   N233 : DINT[1] := ([0] := 9);
   N24 : DINT[31] := ([0] := 100, [1] := 1, [2] := 100, [3] := 1, [4] := 5, [5] := 5, [6] := 60, [7] := 1, [8] := 100, [9] := 1, [10] := 100, [11] := 1, [12] := 5, [13] := 5, [14] := 60, [15] := 1);
   N240 : DINT[68] := ([8] := 254, [10] := -256, [50] := 128, [51] := 9, [52] := 210, [54] := 1, [55] := 210, [60] := 25600, [61] := 9, [62] := 210, [64] := 17408, [66] := 210);
   N241 : DINT[1];
   N242 : DINT[2] := ([0] := -9, [1] := -9);
   N250 : DINT[100] := ([8] := 99, [10] := -256, [50] := -32640, [51] := 9, [52] := 200, [54] := 1, [55] := 200, [61] := 9, [62] := 200, [65] := 1, [66] := 200);
   N251 : DINT[100];
   N252 : DINT[100] := ([0] := -9, [1] := -9);
   N26 : DINT[33] := ([1] := 8, [10] := 38, [11] := 1, [30] := -15194, [31] := 8);
   N27 : DINT[50] := ([40] := 28176, [41] := 29344, [42] := 23976, [43] := 25960, [44] := 29304, [45] := 27664, [46] := 28928, [47] := 16);
   N28 : DINT[17] := ([0] := 124, [1] := 158, [2] := 937, [3] := 50, [4] := 9, [5] := 156, [6] := 3, [10] := 1000, [12] := 100);
   N7 : DINT[100] := ([0] := 5, [1] := 20, [2] := 20, [4] := 30000, [7] := 48, [8] := 48, [9] := 48, [10] := 53, [11] := 53, [12] := 43, [13] := 46, [14] := 46, [15] := 46, [16] := 51, [17] := 51, [18] := 46, [50] := 1, [51] := 1, [52] := 1, [53] := 1, [54] := 1, [55] := 1, [56] := 1, [57] := 1, [58] := 1, [59] := 1, [60] := 1, [61] := 1, [62] := 1, [93] := 9, [99] := 9);
   N_RECVING_PIT_GATE_AUTO : ALIAS FOR Local:0:I.Data.2;
   N_RECVING_PIT_GATE_CLOSE : ALIAS FOR Local:5:O.Data.5;
   N_RECVING_PIT_GATE_OPEN : ALIAS FOR Local:5:O.Data.4;
   NU : DINT;
   O10 : ALIAS FOR R1S0_AENTR:10:O.Data;
   O10_000_Bit00 : ALIAS FOR O10.0;
   O10_000_Bit01 : ALIAS FOR O10.1;
   O10_000_Bit02 : ALIAS FOR O10.2;
   O10_000_Bit03 : ALIAS FOR O10.3;
   O10_000_Bit04 : ALIAS FOR O10.4;
   O10_000_Bit05 : ALIAS FOR O10.5;
   O10_000_Bit06 : ALIAS FOR O10.6;
   O10_000_Bit07 : ALIAS FOR O10.7;
   O10_000_Bit08 : ALIAS FOR O10.8;
   O10_000_Bit09 : ALIAS FOR O10.9;
   O10_000_Bit10 : ALIAS FOR O10.10;
   O10_000_Bit11 : ALIAS FOR O10.11;
   O10_000_Bit12 : ALIAS FOR O10.12;
   O10_000_Bit13 : ALIAS FOR O10.13;
   O10_000_Bit14 : ALIAS FOR O10.14;
   O10_000_Bit15 : ALIAS FOR O10.15;
   O11 : ALIAS FOR R1S0_AENTR:11:O.Data;
   O11_000_Bit00 : ALIAS FOR O11.0;
   O11_000_Bit01 : ALIAS FOR O11.1;
   O11_000_Bit02 : ALIAS FOR O11.2;
   O11_000_Bit03 : ALIAS FOR O11.3;
   O11_000_Bit04 : ALIAS FOR O11.4;
   O11_000_Bit05 : ALIAS FOR O11.5;
   O11_000_Bit06 : ALIAS FOR O11.6;
   O11_000_Bit07 : ALIAS FOR O11.7;
   O11_000_Bit08 : ALIAS FOR O11.8;
   O11_000_Bit09 : ALIAS FOR O11.9;
   O11_000_Bit10 : ALIAS FOR O11.10;
   O11_000_Bit11 : ALIAS FOR O11.11;
   O11_000_Bit12 : ALIAS FOR O11.12;
   O11_000_Bit13 : ALIAS FOR O11.13;
   O11_000_Bit14 : ALIAS FOR O11.14;
   O12 : ALIAS FOR R1S0_AENTR:12:O.Data;
   O12_000_Bit00 : ALIAS FOR O12.0;
   O12_000_Bit01 : ALIAS FOR O12.1;
   O12_000_Bit02 : ALIAS FOR O12.2;
   O12_000_Bit03 : ALIAS FOR O12.3;
   O12_000_Bit04 : ALIAS FOR O12.4;
   O12_000_Bit05 : ALIAS FOR O12.5;
   O12_000_Bit06 : ALIAS FOR O12.6;
   O12_000_Bit08 : ALIAS FOR O12.8;
   O12_000_Bit09 : ALIAS FOR O12.9;
   O12_000_Bit10 : ALIAS FOR O12.10;
   O12_000_Bit11 : ALIAS FOR O12.11;
   O12_000_Bit12 : ALIAS FOR O12.12;
   O12_000_Bit13 : ALIAS FOR O12.13;
   O12_000_Bit14 : ALIAS FOR O12.14;
   O12_000_Bit15 : ALIAS FOR O12.15;
   O13 : ALIAS FOR R2S0_AENTR:1:O.Data;
   O13_000_Bit00 : ALIAS FOR O13.0;
   O13_000_Bit01 : ALIAS FOR O13.1;
   O13_000_Bit02 : ALIAS FOR O13.2;
   O13_000_Bit03 : ALIAS FOR O13.3;
   O13_000_Bit04 : ALIAS FOR O13.4;
   O13_000_Bit05 : ALIAS FOR O13.5;
   O13_000_Bit06 : ALIAS FOR O13.6;
   O13_000_Bit07 : ALIAS FOR O13.7;
   O13_000_Bit08 : ALIAS FOR O13.8;
   O13_000_Bit09 : ALIAS FOR O13.9;
   O13_000_Bit10 : ALIAS FOR O13.10;
   O13_000_Bit15 : ALIAS FOR O13.15;
   O16 : INT[12] := ([0] := 2#0000_1000_0101_1010, [1] := 2#0000_1000_0101_1010, [2] := 2#0000_1000_0101_1010, [3] := 2#0000_1000_0101_1010, [4] := 2#0000_1000_0101_1010, [5] := 2#0000_1000_0101_1010, [6] := 2#0000_1000_0101_1010, [7] := 2#0000_1000_0101_1010);
   O17 : INT[12] := ([0] := 2#0000_1000_0101_1010, [1] := 2#0000_1000_0101_1010, [2] := 2#0000_1000_0101_1010, [3] := 2#0000_1000_0101_1010, [4] := 2#0000_1000_0101_1010, [5] := 2#0000_1000_0101_1010, [6] := 2#0000_1000_0101_1010, [7] := 2#0000_1000_0101_1010);
   O18 : INT[12] := ([0] := 2#0000_1000_0101_1010, [1] := 2#0000_1000_0101_1010, [2] := 2#0000_1000_0101_1010, [3] := 2#0000_1000_0101_1010, [4] := 2#0000_1000_0101_1010, [5] := 2#0000_1000_0101_1010, [6] := 2#0000_1010_1001_1101, [7] := 2#0000_1010_1001_1101);
   O24 : INT[32] := ([7] := 2#0000_0000_1000_0010);
   O24_001_Bit00 : ALIAS FOR O24[1].0;
   O24_001_Bit01 : ALIAS FOR O24[1].1;
   O24_001_Bit02 : ALIAS FOR O24[1].2;
   O24_001_Bit03 : ALIAS FOR O24[1].3;
   O24_001_Bit04 : ALIAS FOR O24[1].4;
   O24_005_Bit00 : ALIAS FOR O24[5].0;
   O24_005_Bit01 : ALIAS FOR O24[5].1;
   O24_005_Bit02 : ALIAS FOR O24[5].2;
   O24_005_Bit03 : ALIAS FOR O24[5].3;
   O24_005_Bit04 : ALIAS FOR O24[5].4;
   O24_005_Bit05 : ALIAS FOR O24[5].5;
   O24_005_Bit06 : ALIAS FOR O24[5].6;
   O24_005_Bit07 : ALIAS FOR O24[5].7;
   O24_005_Bit08 : ALIAS FOR O24[5].8;
   O24_005_Bit09 : ALIAS FOR O24[5].9;
   O24_005_Bit10 : ALIAS FOR O24[5].10;
   O24_005_Bit11 : ALIAS FOR O24[5].11;
   O24_005_Bit12 : ALIAS FOR O24[5].12;
   O24_005_Bit15 : ALIAS FOR O24[5].15;
   O24_007_Bit00 : ALIAS FOR O24[7].0;
   O24_007_Bit01 : ALIAS FOR O24[7].1;
   O24_007_Bit04 : ALIAS FOR O24[7].4;
   O24_007_Bit05 : ALIAS FOR O24[7].5;
   O24_007_Bit06 : ALIAS FOR O24[7].6;
   O24_007_Bit07 : ALIAS FOR O24[7].7;
   O24_007_Bit10 : ALIAS FOR O24[7].10;
   O24_007_Bit11 : ALIAS FOR O24[7].11;
   O24_007_Bit12 : ALIAS FOR O24[7].12;
   O24_007_Bit13 : ALIAS FOR O24[7].13;
   O24_007_Bit14 : ALIAS FOR O24[7].14;
   O24_007_Bit8 : DINT;
   O25 : INT[32] := ([8] := 2#0100_0001_1101_1110, [9] := 2#0011_0111_0100_0010, [10] := 2#1110_0000_0100_0000, [11] := 2#0000_0000_0000_1010);
   O25_008_Bit00 : ALIAS FOR O25[8].0;
   O25_008_Bit01 : ALIAS FOR O25[8].1;
   O25_008_Bit02 : ALIAS FOR O25[8].2;
   O25_008_Bit03 : ALIAS FOR O25[8].3;
   O25_008_Bit04 : ALIAS FOR O25[8].4;
   O25_008_Bit06 : ALIAS FOR O25[8].6;
   O25_008_Bit07 : ALIAS FOR O25[8].7;
   O25_008_Bit08 : ALIAS FOR O25[8].8;
   O25_008_Bit09 : ALIAS FOR O25[8].9;
   O25_008_Bit10 : ALIAS FOR O25[8].10;
   O25_008_Bit12 : ALIAS FOR O25[8].12;
   O25_008_Bit13 : ALIAS FOR O25[8].13;
   O25_008_Bit14 : ALIAS FOR O25[8].14;
   O25_008_Bit15 : ALIAS FOR O25[8].15;
   O25_009_Bit00 : ALIAS FOR O25[9].0;
   O25_009_Bit01 : ALIAS FOR O25[9].1;
   O25_009_Bit02 : ALIAS FOR O25[9].2;
   O25_009_Bit03 : ALIAS FOR O25[9].3;
   O25_009_Bit04 : ALIAS FOR O25[9].4;
   O25_009_Bit05 : ALIAS FOR O25[9].5;
   O25_009_Bit06 : ALIAS FOR O25[9].6;
   O25_009_Bit07 : ALIAS FOR O25[9].7;
   O25_009_Bit08 : ALIAS FOR O25[9].8;
   O25_009_Bit09 : ALIAS FOR O25[9].9;
   O25_009_Bit10 : ALIAS FOR O25[9].10;
   O25_009_Bit11 : ALIAS FOR O25[9].11;
   O25_009_Bit12 : ALIAS FOR O25[9].12;
   O25_009_Bit13 : ALIAS FOR O25[9].13;
   O25_009_Bit14 : ALIAS FOR O25[9].14;
   O25_009_Bit15 : ALIAS FOR O25[9].15;
   O25_010_Bit00 : ALIAS FOR O25[10].0;
   O25_010_Bit01 : ALIAS FOR O25[10].1;
   O25_010_Bit02 : ALIAS FOR O25[10].2;
   O25_010_Bit03 : ALIAS FOR O25[10].3;
   O25_010_Bit04 : ALIAS FOR O25[10].4;
   O25_010_Bit05 : ALIAS FOR O25[10].5;
   O25_010_Bit06 : ALIAS FOR O25[10].6;
   O25_010_Bit07 : ALIAS FOR O25[10].7;
   O25_010_Bit08 : ALIAS FOR O25[10].8;
   O25_010_Bit09 : ALIAS FOR O25[10].9;
   O25_010_Bit10 : ALIAS FOR O25[10].10;
   O25_010_Bit11 : ALIAS FOR O25[10].11;
   O25_010_Bit12 : ALIAS FOR O25[10].12;
   O25_010_Bit13 : ALIAS FOR O25[10].13;
   O25_010_Bit14 : ALIAS FOR O25[10].14;
   O25_010_Bit15 : ALIAS FOR O25[10].15;
   O25_011_Bit00 : ALIAS FOR O25[11].0;
   O25_011_Bit01 : ALIAS FOR O25[11].1;
   O25_011_Bit03 : ALIAS FOR O25[11].3;
   O25_011_Bit14 : ALIAS FOR O25[11].14;
   O25_011_Bit15 : ALIAS FOR O25[11].15;
   O25_012_Bit00 : ALIAS FOR O25[12].0;
   O25_012_Bit01 : ALIAS FOR O25[12].1;
   O25_012_Bit02 : ALIAS FOR O25[12].2;
   O25_012_Bit03 : ALIAS FOR O25[12].3;
   O25_012_Bit04 : ALIAS FOR O25[12].4;
   O25_012_Bit05 : ALIAS FOR O25[12].5;
   O25_012_Bit06 : ALIAS FOR O25[12].6;
   O25_012_Bit07 : ALIAS FOR O25[12].7;
   O25_012_Bit08 : ALIAS FOR O25[12].8;
   O25_012_Bit09 : ALIAS FOR O25[12].9;
   O25_012_Bit10 : ALIAS FOR O25[12].10;
   O25_012_Bit11 : ALIAS FOR O25[12].11;
   O25_012_Bit12 : ALIAS FOR O25[12].12;
   O25_012_Bit13 : ALIAS FOR O25[12].13;
   O25_012_Bit14 : ALIAS FOR O25[12].14;
   O9 : ALIAS FOR R1S0_AENTR:9:O.Data;
   O9_000_Bit00 : ALIAS FOR O9.0;
   O9_000_Bit01 : ALIAS FOR O9.1;
   O9_000_Bit02 : ALIAS FOR O9.2;
   O9_000_Bit03 : ALIAS FOR O9.3;
   O9_000_Bit04 : ALIAS FOR O9.4;
   O9_000_Bit05 : ALIAS FOR O9.5;
   O9_000_Bit06 : ALIAS FOR O9.6;
   O9_000_Bit07 : ALIAS FOR O9.7;
   O9_000_Bit08 : ALIAS FOR O9.8;
   O9_000_Bit09 : ALIAS FOR O9.9;
   O9_000_Bit10 : ALIAS FOR O9.10;
   O9_000_Bit11 : ALIAS FOR O9.11;
   O9_000_Bit12 : ALIAS FOR O9.12;
   O9_000_Bit13 : ALIAS FOR O9.13;
   O9_000_Bit14 : ALIAS FOR O9.14;
   O9_000_Bit15 : ALIAS FOR O9.15;
   OLIVER_BIN : ALIAS FOR I4.8;
   OLIVER_SEP : ALIAS FOR I25[3].11;
   output_Bit : BOOL;
   Output_Bit_2 : BOOL;
   P10_ALARM : ALIAS FOR T4[97];
   P10_ALARM1 : ALIAS FOR T4[99];
   P10_AUTO_S : ALIAS FOR B3[5].10;
   P10_FLOW_A : ALIAS FOR N13[82];
   P10_FLOW_P : ALIAS FOR I24[21].8;
   P10_FLOW_P1 : ALIAS FOR C5[39];
   P10_FLW_OZ : ALIAS FOR N13[80];
   P10_MB : ALIAS FOR B12[10].2;
   P10_NO_FLO : ALIAS FOR B12[10].3;
   P10_OZ : ALIAS FOR N13[81];
   P10_RUN_AU : ALIAS FOR O24[5].9;
   P10_RUN_AU1 : ALIAS FOR B3[4].10;
   P10_SEC_SE : ALIAS FOR B17[1].10;
   P10_SEL_SW : ALIAS FOR I24[4].9;
   P10_SET : ALIAS FOR B12[10].0;
   P10_SPEED : ALIAS FOR N13[84];
   P10_STOP : ALIAS FOR B12[10].1;
   P11_RUN_AU : ALIAS FOR O24[5].10;
   P11_SEL_SW : ALIAS FOR I24[4].10;
   P12_RUN_AU : ALIAS FOR O24[5].11;
   P12_SEL_SW : ALIAS FOR I24[4].11;
   P1_ALARM_N : ALIAS FOR T4[81];
   P1_ALARM_N1 : ALIAS FOR T4[82];
   P1_AUTO_SE : ALIAS FOR B3[5].1;
   P1_FLOW_AN : ALIAS FOR N13[2];
   P1_FLOW_PL : ALIAS FOR C5[30];
   P1_FLOW_PU : ALIAS FOR I24[21].0;
   P1_FLW_OZ : ALIAS FOR N13[0];
   P1_MB : ALIAS FOR B12[1].2;
   P1_NO_FLOW : ALIAS FOR B12[1].3;
   P1_OZ : ALIAS FOR N13[1];
   P1_RUN_AUT : ALIAS FOR O24[5].0;
   P1_RUN_AUT1 : ALIAS FOR B3[4].1;
   P1_SEC_SEL : ALIAS FOR B17[1].1;
   P1_SEL_SW : ALIAS FOR I24[4].0;
   P1_SET : ALIAS FOR B12[1].0;
   P1_SPEED_O : ALIAS FOR N13[4];
   P1_STOP : ALIAS FOR B12[1].1;
   P2_ALARM_N : ALIAS FOR T4[83];
   P2_ALARM_N1 : ALIAS FOR T4[84];
   P2_AUTO_SE : ALIAS FOR B3[5].2;
   P2_FLOW_AN : ALIAS FOR N13[12];
   P2_FLOW_PL : ALIAS FOR C5[32];
   P2_FLOW_PU : ALIAS FOR I24[21].1;
   P2_FLW_OZ : ALIAS FOR N13[10];
   P2_MB : ALIAS FOR B12[2].2;
   P2_NO_FLOW : ALIAS FOR B12[2].3;
   P2_OZ : ALIAS FOR N13[11];
   P2_RUN_AUT : ALIAS FOR O24[5].1;
   P2_RUN_AUT1 : ALIAS FOR B3[4].2;
   P2_SEC_SEL : ALIAS FOR B17[1].2;
   P2_SEL_SW : ALIAS FOR I24[4].1;
   P2_SET : ALIAS FOR B12[2].0;
   P2_SPEED_O : ALIAS FOR N13[14];
   P2_STOP : ALIAS FOR B12[2].1;
   P3_ALARM_N : ALIAS FOR T4[85];
   P3_ALARM_N1 : ALIAS FOR T4[86];
   P3_AUTO_SE : ALIAS FOR B3[5].3;
   P3_FLOW_AN : ALIAS FOR N13[22];
   P3_FLOW_PL : ALIAS FOR C5[33];
   P3_FLOW_PU : ALIAS FOR I24[21].2;
   P3_FLW_OZ : ALIAS FOR N13[20];
   P3_MB : ALIAS FOR B12[3].2;
   P3_NO_FLOW : ALIAS FOR B12[3].3;
   P3_OZ : ALIAS FOR N13[21];
   P3_RUN_AUT : ALIAS FOR O24[5].2;
   P3_RUN_AUT1 : ALIAS FOR B3[4].3;
   P3_SEC_SEL : ALIAS FOR B17[1].3;
   P3_SEL_SW : ALIAS FOR I24[4].2;
   P3_SET : ALIAS FOR B12[3].0;
   P3_SPEED_O : ALIAS FOR N13[24];
   P3_STOP : ALIAS FOR B12[3].1;
   P4_ALARM_N : ALIAS FOR T4[87];
   P4_ALARM_N1 : ALIAS FOR T4[88];
   P4_AUTO_SE : ALIAS FOR B3[5].4;
   P4_FLOW_AN : ALIAS FOR N13[32];
   P4_FLOW_PL : ALIAS FOR C5[34];
   P4_FLOW_PU : ALIAS FOR I24[21].3;
   P4_FLW_OZ : ALIAS FOR N13[30];
   P4_MB : ALIAS FOR B12[4].2;
   P4_NO_FLOW : ALIAS FOR B12[4].3;
   P4_OZ : ALIAS FOR N13[31];
   P4_RUN_AUT : ALIAS FOR O24[5].3;
   P4_RUN_AUT1 : ALIAS FOR B3[4].4;
   P4_SEC_SEL : ALIAS FOR B17[1].4;
   P4_SEL_SW : ALIAS FOR I24[4].3;
   P4_SET : ALIAS FOR B12[4].0;
   P4_SPEED_O : ALIAS FOR N13[34];
   P4_STOP : ALIAS FOR B12[4].1;
   P5_ALARM_N : ALIAS FOR T4[89];
   P5_ALARM_N1 : ALIAS FOR T4[90];
   P5_AUTO_SE : ALIAS FOR B3[5].5;
   P5_FLOW_AN : ALIAS FOR N13[42];
   P5_FLOW_PL : ALIAS FOR C5[35];
   P5_FLOW_PU : ALIAS FOR I24[21].4;
   P5_FLW_OZ : ALIAS FOR N13[40];
   P5_MB : ALIAS FOR B12[5].2;
   P5_NO_FLOW : ALIAS FOR B12[5].3;
   P5_OZ : ALIAS FOR N13[41];
   P5_RUN_AUT : ALIAS FOR O24[5].4;
   P5_RUN_AUT1 : ALIAS FOR B3[4].5;
   P5_SEC_SEL : ALIAS FOR B17[1].5;
   P5_SEL_SW : ALIAS FOR I24[4].4;
   P5_SET : ALIAS FOR B12[5].0;
   P5_SPEED_O : ALIAS FOR N13[44];
   P5_STOP : ALIAS FOR B12[5].1;
   P6_ALARM_N : ALIAS FOR T4[91];
   P6_ALARM_N1 : ALIAS FOR T4[92];
   P6_AUTO_SE : ALIAS FOR B3[5].6;
   P6_FLOW_AN : ALIAS FOR N13[52];
   P6_FLOW_PL : ALIAS FOR C5[36];
   P6_FLOW_PU : ALIAS FOR I24[21].5;
   P6_FLW_OZ : ALIAS FOR N13[50];
   P6_MB : ALIAS FOR B12[6].2;
   P6_NO_FLOW : ALIAS FOR B12[6].3;
   P6_OZ : ALIAS FOR N13[51];
   P6_RUN_AUT : ALIAS FOR O24[5].5;
   P6_RUN_AUT1 : ALIAS FOR B3[4].6;
   P6_SEC_SEL : ALIAS FOR B17[1].6;
   P6_SEL_SW : ALIAS FOR I24[4].5;
   P6_SET : ALIAS FOR B12[6].0;
   P6_SPEED_O : ALIAS FOR N13[54];
   P6_STOP : ALIAS FOR B12[6].1;
   P7_ALARM_N : ALIAS FOR T4[93];
   P7_ALARM_N1 : ALIAS FOR T4[94];
   P7_AUTO_SE : ALIAS FOR B3[5].7;
   P7_FLOW_AN : ALIAS FOR N13[62];
   P7_FLOW_PL : ALIAS FOR C5[37];
   P7_FLOW_PU : ALIAS FOR I24[21].6;
   P7_FLW_OZ : ALIAS FOR N13[60];
   P7_MB : ALIAS FOR B12[7].2;
   P7_NO_FLOW : ALIAS FOR B12[7].3;
   P7_OZ : ALIAS FOR N13[61];
   P7_RUN_AUT : ALIAS FOR O24[5].6;
   P7_RUN_AUT1 : ALIAS FOR B3[4].7;
   P7_SEC_SEL : ALIAS FOR B17[1].7;
   P7_SEL_SW : ALIAS FOR I24[4].6;
   P7_SET : ALIAS FOR B12[7].0;
   P7_SPEED_O : ALIAS FOR N13[64];
   P7_STOP : ALIAS FOR B12[7].1;
   P8_ALARM_N : ALIAS FOR T4[95];
   P8_ALARM_N1 : ALIAS FOR T4[96];
   P8_AUTO_SE : ALIAS FOR B3[5].8;
   P8_FLOW_AN : ALIAS FOR N13[72];
   P8_FLOW_PL : ALIAS FOR C5[38];
   P8_FLOW_PU : ALIAS FOR I24[21].7;
   P8_FLW_OZ : ALIAS FOR N13[70];
   P8_MB : ALIAS FOR B12[8].2;
   P8_NO_FLOW : ALIAS FOR B12[8].3;
   P8_OZ : ALIAS FOR N13[71];
   P8_RUN_AUT : ALIAS FOR O24[5].7;
   P8_RUN_AUT1 : ALIAS FOR B3[4].8;
   P8_SEC_SEL : ALIAS FOR B17[1].8;
   P8_SEL_SW : ALIAS FOR I24[4].7;
   P8_SET : ALIAS FOR B12[8].0;
   P8_SPEED_O : ALIAS FOR N13[74];
   P8_STOP : ALIAS FOR B12[8].1;
   P9_RUN_AUT : ALIAS FOR O24[5].8;
   P9_SEC_SEL : ALIAS FOR B17[1].9;
   P9_SEL_SW : ALIAS FOR I24[4].8;
   P_RESET_AU : ALIAS FOR B3[4].0;
   PMP_15_OFF_DLY : REAL := 5.0;
   PMP_15_OFF_DLY_SCALE : REAL := 5000.0;
   PMP_15_ON_DLY : REAL := 5.0;
   PMP_15_ON_DLY_SCALE : REAL := 5000.0;
   PMP_15_TMR : TIMER := (PRE := 5000);
   PMP_15_TMR_2 : TIMER := (PRE := 5000);
   ProcessAll : BOOL;
   PUMP_13_RUN : ALIAS FOR R3M1_AENTR:3:O.8;
   PUMP_14_RUN : ALIAS FOR R3M1_AENTR:3:O.9;
   PUMP_15_AUTO : BOOL;
   PUMP_15_RUN : ALIAS FOR R3M1_AENTR:3:O.14;
   PUMP_NO_FL : ALIAS FOR B12[11].0;
   R6 : CONTROL[1];
   Rack24_1_Mode : BOOL := 1;
   RemoteAndcoAnalogIn : DINT[40] := ([1] := 9993, [3] := 10270, [4] := 5041, [5] := 7694, [7] := 9661, [9] := 3611, [10] := 9885, [11] := 8109, [12] := 10717, [13] := 7657, [14] := 9078, [15] := 8853, [19] := 9087, [20] := 9586);
   RSSql_MSG_BTR : INT;
   RSSql_MSG_BTR_DN : ALIAS FOR RSSql_MSG_BTR.0;
   RSSql_MSG_BTR_ER : ALIAS FOR RSSql_MSG_BTR.1;
   RSSql_MSG_Control : MESSAGE;
        MessageParameters(ServiceCode := 16#004d, LocalElement := spTicketTableBay1Wt, ...)
   RSSql_MSG_Data : DINT := 138;
   RSSql_MSG_En : BOOL;
   RSVIEW_ALA : ALIAS FOR B3[0].11;
   S : INT[83] := ([0] := 16#0004, [1] := 16#00de, [2] := 16#9032, [3] := 16#a005, [4] := 16#455e, [5] := 16#4000, [9] := 16#0002, [10] := 16#0032, [11] := 16#ffff, [12] := 16#ffff, [17] := 16#0002, [20] := 16#0001, [21] := 16#0008, [22] := 16#0006, [23] := 16#0005, [27] := 16#ffff, [28] := 16#ffff, [33] := 16#0208, [35] := 16#0030, [54] := 16#0021, [57] := 16#01f5, [58] := 16#0002, [59] := 16#0006, [60] := 16#0227, [61] := 16#0001, [62] := 16#0004, [63] := 16#0801, [64] := 16#0005, [65] := 16#0010, [66] := 16#0200);
   S24 : ALIAS FOR S[24];
   SCP_AOI : SCP_Inv[8] := ([0].In := 28184.0, [0].InRawMin := 12336.0, [0].InRawMax := 28816.0, [0].InEUMax := 3200.0, [0].Out := 122.71826, [1].In := 29344.0, [1].InRawMin := 10744.0, [1].InRawMax := 30320.0, [1].InEUMax := 3200.0, [1].Out := 159.54224, [2].In := 23976.0, [2].InRawMin := 9280.0, [2].InRawMax := 30064.0, [2].InEUMax := 3200.0, [2].Out := 937.3364, [3].In := 25960.0, [3].InRawMin := 7368.0, [3].InRawMax := 26256.0, [3].InEUMax := 3200.0, [3].Out := 50.148193, [4].In := 29296.0, [4].InRawMin := 9080.0, [4].InRawMax := 29360.0, [4].InEUMax := 3200.0, [4].Out := 10.098633, [5].In := 27664.0, [5].InRawMin := 8256.0, [5].InRawMax := 28656.0, [5].InEUMax := 3200.0, [5].Out := 155.60791, [6].In := 28928.0, [6].InRawMin := 11696.0, [6].InRawMax := 28944.0, [6].InEUMax := 3200.0, [6].Out := 2.9685059);
   Screen_Cancel : DINT;
   SCREENER_DRAG_START : BOOL;
   SCREENER_DRAG_STOP : BOOL;
   SCREENER_LEG_START : BOOL;
   SCREENER_LEG_STOP : BOOL;
   SCREENINGS : ALIAS FOR I7.15;
   Select_Cal_Bins : BOOL;
   Select_Clean_Bins : BOOL := 1;
   Select_Treat_Bins : BOOL;
   sendData : BOOL;
   sendData1 : BOOL;
   sendData_ONS : DINT;
   spBinGateRates : DINT[50] := ([11] := 86, [12] := 95, [13] := 79, [14] := 94, [15] := 93, [16] := 31, [17] := 79, [21] := 95, [22] := 83, [23] := 97, [24] := 90, [25] := 103, [26] := 99);
   spCapGrossWt : BOOL;
   spCapTareWt : BOOL;
   spCreateTicket : BOOL;
   spShowCreateTicketPB : BOOL;
   spTicketBinActive : DINT;
   spTicketBinSet : DINT;
   spTicketProcessing : BOOL;
   spTicketProcessStr : BOOL;
   spTicketTableBay1GrsWt : DINT;
   spTicketTableBay1Wt : DINT;
   spVAR_BINARRAY : STRING[50] := ([11] := '803001-Azimut-Certified - Limagrain  - HRW Seed Wheat', [12] := '883004-Lenetah-Certified -   - Barley Seed', [15] := '843002-Expresso-Certified-Monsanto -DNS Seed Wheat', [16] := '843005-Glee -Certified-WSU -DNS Seed Wheat', [17] := '843006-Kelse-Certified-WSU -DNS Seed Wheat', [22] := '843001-Buck Pronto-Certified-Limagrain -DNS Seed Wheat', [23] := '843004-SY 605-Certified-Sygenta Clearfield-DNS Seed Wheat', [24] := '803004-Keldin -Certified-Monsanto -HRW Seed Wheat', [25] := '843001-Buck Pronto-Certified-Limagrain -DNS Seed Wheat', [26] := '843003-Solano-Certified - Monsanto  - DNS Seed Wheat');
   sqlIndex : DINT;
   sqlIndex1 : DINT;
   sqlNewStartWeight : BOOL;
   sqlNewTreatment : BOOL;
   sqlNewTreatments_ONS : DINT;
   sqlNewVariety : BOOL;
   sqlNewVariety_ONS : DINT;
   sqlStartWtRecvd : DINT := 1;
   sqlTreatID : DINT;
   sqlTreatmentsRevd : DINT;
   sqlTreatRate : DINT;
   sqlTrtSendDelayTMR : TIMER := (PRE := 1000);
   sqlVaritiesRevd : DINT;
   sqlVarityID : DINT;
   sqlVarityRate : DINT;
   sqlVarSendDelayTMR : TIMER := (PRE := 1000);
   strEmptyVar : STRING := 'Empty';
   SURGE_BIN_HI : ALIAS FOR Local:0:I.Data.0;
   SURGE_BIN_LO : ALIAS FOR Local:0:I.Data.1;
   SWW_Index : DINT := 100;
   SWW_Variety_DB : Varieties_DB[100] := ([0].Id := 821001, [0].Name := 'ArtDeco', [0].ClassId := 1, [0].ClassType := 'Foundation', [0].MarketClassId := 82, [0].MarketClassType := 'SWW', [0].FullDecription := '821001  ArtDeco  Foundation  SWW', [1].Id := 822001, [1].Name := 'ArtDeco', [1].ClassId := 2, [1].ClassType := 'Registered', [1].MarketClassId := 82, [1].MarketClassType := 'SWW', [1].FullDecription := '822001  ArtDeco  Registered  SWW', [2].Id := 823001, [2].Name := 'ArtDeco', [2].ClassId := 3, [2].ClassType := 'Certified', [2].MarketClassId := 82, [2].MarketClassType := 'SWW', [2].FullDecription := '823001  ArtDeco  Certified  SWW', [3].Id := 821002, [3].Name := 'Huffman', [3].ClassId := 1, [3].ClassType := 'Foundation', [3].MarketClassId := 82, [3].MarketClassType := 'SWW', [3].FullDecription := '821002  Huffman  Foundation  SWW', [4].Id := 822002, [4].Name := 'Huffman', [4].ClassId := 2, [4].ClassType := 'Registered', [4].MarketClassId := 82, [4].MarketClassType := 'SWW', [4].FullDecription := '822002  Huffman  Registered  SWW', [5].Id := 823002, [5].Name := 'Huffman', [5].ClassId := 3, [5].ClassType := 'Certified', [5].MarketClassId := 82, [5].MarketClassType := 'SWW', [5].FullDecription := '823002  Huffman  Certified  SWW', [6].Id := 821003, [6].Name := 'WB 1035 CL Spring', [6].ClassId := 1, [6].ClassType := 'Foundation', [6].MarketClassId := 82, [6].MarketClassType := 'SWW', [6].FullDecription := '821003  WB 1035 CL Spring Foundation  SWW', [7].Id := 822003, [7].Name := 'WB 1035 CL Spring', [7].ClassId := 2, [7].ClassType := 'Registered', [7].MarketClassId := 82, [7].MarketClassType := 'SWW', [7].FullDecription := '822003  WB 1035 CL Spring  Registered  SWW', [8].Id := 823003, [8].Name := 'WB 1035 CL Spring', [8].ClassId := 3, [8].ClassType := 'Certified',
        [8].MarketClassId := 82, [8].MarketClassType := 'SWW', [8].FullDecription := '823003  WB 1035 CL Spring  Certified SWW');
   SWW_VarietySize : DINT := 100;
   SYMBOL : ALIAS FOR B3[0].0;
   SYMBOL_ANA : ALIAS FOR N10[1];
   T11 : TIMER[100] := ([0].PRE := 500, [0].ACC := 500, [0].EN := 1, [0].DN := 1, [1].PRE := 500, [1].ACC := 125, [1].EN := 1, [1].TT := 1, [3].PRE := 600000, [4].PRE := 1000, [5].PRE := 5000, [6].PRE := 5000, [7].PRE := 600000, [10].PRE := 5000, [11].PRE := 5000, [12].PRE := 5000, [13].PRE := 5000, [14].PRE := 5000, [15].PRE := 25000, [16].PRE := 5000, [17].PRE := 5000, [18].PRE := 5000, [19].PRE := 20000, [19].ACC := 20000, [19].EN := 1, [19].DN := 1);
   T11_AIR_SV : ALIAS FOR O9.0;
   T11_AIRSG : ALIAS FOR I1.0;
   T11_AIRSG1 : ALIAS FOR T4[0];
   T11_AIRSG2 : ALIAS FOR T4[1];
   T11_ASCII : ALIAS FOR B17[11].1;
   T11_ASSII : ALIAS FOR A16[112];
   T11_ASSII1 : ALIAS FOR A16[115];
   T11_AUTO_A : ALIAS FOR T4[61];
   T11_AUTO_A1 : ALIAS FOR T4[61].PRE;
   T11_AUTO_A2 : ALIAS FOR T4[61].ACC;
   T11_AUTO_M : ALIAS FOR B3[11].1;
   T11_AUTO_S : ALIAS FOR B3[11].14;
   T11_BINDIC : ALIAS FOR I4.11;
   T11_CAL_CL : ALIAS FOR B15[51].3;
   T11_CAL_LA : ALIAS FOR B15[51].2;
   T11_CAL_OP : ALIAS FOR B15[51].4;
   T11_CAL_ST : ALIAS FOR B15[51].1;
   T11_CLOSE : ALIAS FOR O9.1;
   T11_CLOSE1 : ALIAS FOR B3[11].9;
   T11_CLOSE2 : ALIAS FOR B3[11].11;
   T11_CORREC : ALIAS FOR F8[2];
   T11_DLY_TR : ALIAS FOR T4[0].PRE;
   T11_DLY_TR1 : ALIAS FOR T4[0].ACC;
   T11_DLY_TR2 : ALIAS FOR T4[1].PRE;
   T11_DLY_TR3 : ALIAS FOR T4[1].ACC;
   T11_FAULT : ALIAS FOR B3[11].15;
   T11_GATE_C : ALIAS FOR C5[11];
   T11_GATE_C1 : ALIAS FOR C5[11].PRE;
   T11_GATE_C2 : ALIAS FOR C5[11].ACC;
   T11_HOLD_A : ALIAS FOR B3[11].3;
   T11_HOLD_M : ALIAS FOR B3[11].6;
   T11_K_FACT : ALIAS FOR F8[1];
   T11_LOW_BI : ALIAS FOR B15[11].2;
   T11_MTR_GT : ALIAS FOR I1.2;
   T11_NO_PAS : ALIAS FOR B17[11].2;
   T11_NULL_V : ALIAS FOR A16[118];
   T11_NULL_V1 : ALIAS FOR A16[119];
   T11_OP_DEF : ALIAS FOR A16[116];
   T11_OP_DEF1 : ALIAS FOR A16[117];
   T11_OP_NAM : ALIAS FOR A16[113];
   T11_OP_NAM1 : ALIAS FOR A16[114];
   T11_OPEN_A : ALIAS FOR B3[11].8;
   T11_OPEN_M : ALIAS FOR O9.2;
   T11_OPEN_M1 : ALIAS FOR B3[11].10;
   T11_RELEAS : ALIAS FOR B3[11].5;
   T11_RESET : ALIAS FOR B3[11].7;
   T11_SET_AU : ALIAS FOR B3[11].2;
   T11_SET_DE : ALIAS FOR B3[2].0;
   T11_SET_LO : ALIAS FOR B3[11].13;
   T11_SET_MA : ALIAS FOR B3[11].12;
   T11_SET_NA : ALIAS FOR A16[110];
   T11_SET_NA1 : ALIAS FOR A16[111];
   T11_SET_NA2 : ALIAS FOR B17[11].0;
   T11_STOP_A : ALIAS FOR B3[11].4;
   T11_TREAT : ALIAS FOR B3[11].0;
   T11_TRT_MO : ALIAS FOR T4[41];
   T11_TRT_MO1 : ALIAS FOR T4[41].PRE;
   T11_TRT_MO2 : ALIAS FOR T4[41].ACC;
   T12_AIR_GA : ALIAS FOR I1.3;
   T12_AIR_SV : ALIAS FOR O9.3;
   T12_ASCII : ALIAS FOR B17[12].1;
   T12_ASSII : ALIAS FOR A16[122];
   T12_ASSII1 : ALIAS FOR A16[125];
   T12_AUTO_A : ALIAS FOR T4[62];
   T12_AUTO_A1 : ALIAS FOR T4[62].PRE;
   T12_AUTO_A2 : ALIAS FOR T4[62].ACC;
   T12_AUTO_M : ALIAS FOR B3[12].1;
   T12_AUTO_S : ALIAS FOR B3[12].14;
   T12_BINDIC : ALIAS FOR I4.12;
   T12_CAL_CL : ALIAS FOR B15[52].3;
   T12_CAL_LA : ALIAS FOR B15[52].2;
   T12_CAL_OP : ALIAS FOR B15[52].4;
   T12_CAL_ST : ALIAS FOR B15[52].1;
   T12_CLOSE : ALIAS FOR O9.4;
   T12_CLOSE1 : ALIAS FOR B3[12].9;
   T12_CLOSE2 : ALIAS FOR B3[12].11;
   T12_CORREC : ALIAS FOR F8[4];
   T12_DLY_TR : ALIAS FOR T4[2];
   T12_DLY_TR1 : ALIAS FOR T4[2].PRE;
   T12_DLY_TR2 : ALIAS FOR T4[2].ACC;
   T12_DLY_TR3 : ALIAS FOR T4[3];
   T12_DLY_TR4 : ALIAS FOR T4[3].PRE;
   T12_DLY_TR5 : ALIAS FOR T4[3].ACC;
   T12_FAULT : ALIAS FOR B3[12].15;
   T12_GATE_C : ALIAS FOR C5[12];
   T12_GATE_C1 : ALIAS FOR C5[12].PRE;
   T12_GATE_C2 : ALIAS FOR C5[12].ACC;
   T12_HOLD_A : ALIAS FOR B3[12].3;
   T12_HOLD_M : ALIAS FOR B3[12].6;
   T12_K_FACT : ALIAS FOR F8[3];
   T12_LOW_BI : ALIAS FOR B15[12].2;
   T12_METER : ALIAS FOR I1.5;
   T12_NO_PAS : ALIAS FOR B17[12].2;
   T12_NULL_V : ALIAS FOR A16[128];
   T12_NULL_V1 : ALIAS FOR A16[129];
   T12_OP_DEF : ALIAS FOR A16[126];
   T12_OP_DEF1 : ALIAS FOR A16[127];
   T12_OP_NAM : ALIAS FOR A16[123];
   T12_OP_NAM1 : ALIAS FOR A16[124];
   T12_OPEN_A : ALIAS FOR B3[12].8;
   T12_OPEN_M : ALIAS FOR O9.5;
   T12_OPEN_M1 : ALIAS FOR B3[12].10;
   T12_RELEAS : ALIAS FOR B3[12].5;
   T12_RESET : ALIAS FOR B3[12].7;
   T12_SET_AU : ALIAS FOR B3[12].2;
   T12_SET_DE : ALIAS FOR B3[2].1;
   T12_SET_LO : ALIAS FOR B3[12].13;
   T12_SET_MA : ALIAS FOR B3[12].12;
   T12_SET_NA : ALIAS FOR A16[120];
   T12_SET_NA1 : ALIAS FOR A16[121];
   T12_SET_NA2 : ALIAS FOR B17[12].0;
   T12_STOP_A : ALIAS FOR B3[12].4;
   T12_TREAT : ALIAS FOR B3[12].0;
   T12_TRT_MO : ALIAS FOR T4[42];
   T12_TRT_MO1 : ALIAS FOR T4[42].PRE;
   T12_TRT_MO2 : ALIAS FOR T4[42].ACC;
   T13_AIR_GA : ALIAS FOR I1.6;
   T13_AIR_SV : ALIAS FOR O9.6;
   T13_ASCII : ALIAS FOR B17[13].1;
   T13_ASSII : ALIAS FOR A16[132];
   T13_ASSII1 : ALIAS FOR A16[135];
   T13_AUTO_A : ALIAS FOR T4[63];
   T13_AUTO_A1 : ALIAS FOR T4[63].PRE;
   T13_AUTO_A2 : ALIAS FOR T4[63].ACC;
   T13_AUTO_M : ALIAS FOR B3[13].1;
   T13_AUTO_S : ALIAS FOR B3[13].14;
   T13_BINDIC : ALIAS FOR I4.13;
   T13_CAL_CL : ALIAS FOR B15[53].3;
   T13_CAL_LA : ALIAS FOR B15[53].2;
   T13_CAL_OP : ALIAS FOR B15[53].4;
   T13_CAL_ST : ALIAS FOR B15[53].1;
   T13_CLOSE : ALIAS FOR O9.7;
   T13_CLOSE1 : ALIAS FOR B3[13].9;
   T13_CLOSE2 : ALIAS FOR B3[13].11;
   T13_CORREC : ALIAS FOR F8[6];
   T13_DLY_TR : ALIAS FOR T4[4];
   T13_DLY_TR1 : ALIAS FOR T4[4].PRE;
   T13_DLY_TR2 : ALIAS FOR T4[4].ACC;
   T13_DLY_TR3 : ALIAS FOR T4[5];
   T13_DLY_TR4 : ALIAS FOR T4[5].PRE;
   T13_DLY_TR5 : ALIAS FOR T4[5].ACC;
   T13_FAULT : ALIAS FOR B3[13].15;
   T13_GATE_C : ALIAS FOR C5[13];
   T13_GATE_C1 : ALIAS FOR C5[13].PRE;
   T13_GATE_C2 : ALIAS FOR C5[13].ACC;
   T13_HOLD_A : ALIAS FOR B3[13].3;
   T13_HOLD_M : ALIAS FOR B3[13].6;
   T13_K_FACT : ALIAS FOR F8[5];
   T13_LOW_BI : ALIAS FOR B15[13].2;
   T13_MTR_GA : ALIAS FOR I1.8;
   T13_NO_PAS : ALIAS FOR B17[13].2;
   T13_NULL_V : ALIAS FOR A16[138];
   T13_NULL_V1 : ALIAS FOR A16[139];
   T13_OP_DEF : ALIAS FOR A16[136];
   T13_OP_DEF1 : ALIAS FOR A16[137];
   T13_OP_NAM : ALIAS FOR A16[133];
   T13_OP_NAM1 : ALIAS FOR A16[134];
   T13_OPEN_A : ALIAS FOR B3[13].8;
   T13_OPEN_M : ALIAS FOR O9.8;
   T13_OPEN_M1 : ALIAS FOR B3[13].10;
   T13_RELEAS : ALIAS FOR B3[13].5;
   T13_RESET : ALIAS FOR B3[13].7;
   T13_SET_AU : ALIAS FOR B3[13].2;
   T13_SET_DE : ALIAS FOR B3[2].2;
   T13_SET_LO : ALIAS FOR B3[13].13;
   T13_SET_MA : ALIAS FOR B3[13].12;
   T13_SET_NA : ALIAS FOR A16[130];
   T13_SET_NA1 : ALIAS FOR A16[131];
   T13_SET_NA2 : ALIAS FOR B17[13].0;
   T13_STOP_A : ALIAS FOR B3[13].4;
   T13_TREAT : ALIAS FOR B3[13].0;
   T13_TRT_MO : ALIAS FOR T4[43];
   T13_TRT_MO1 : ALIAS FOR T4[43].PRE;
   T13_TRT_MO2 : ALIAS FOR T4[43].ACC;
   T13C_AIR_G : ALIAS FOR O12.10;
   T13C_CLOSE : ALIAS FOR T22[6];
   T13C_CLOSE1 : ALIAS FOR T22[6].PRE;
   T13C_CLOSE2 : ALIAS FOR T22[6].ACC;
   T13C_GATE : ALIAS FOR B21[0].0;
   T13C_GATE1 : ALIAS FOR B21[0].1;
   T13C_GATE2 : ALIAS FOR B21[0].3;
   T13C_GATE3 : ALIAS FOR B21[0].4;
   T13C_GATE4 : ALIAS FOR B21[0].5;
   T13C_GATE5 : ALIAS FOR B21[0].6;
   T13C_GATE6 : ALIAS FOR B21[0].7;
   T13C_GATE7 : ALIAS FOR B21[0].8;
   T13C_GATE8 : ALIAS FOR B21[0].9;
   T13C_GATEC : ALIAS FOR B21[0].2;
   T13C_GATET : ALIAS FOR C5[2];
   T13C_SET_D : ALIAS FOR B21[70].14;
   T13C_TMR_A : ALIAS FOR C5[2].ACC;
   T13C_TMR_P : ALIAS FOR C5[2].PRE;
   T13C_TREAT : ALIAS FOR B21[70].10;
   T13C_TRT_M : ALIAS FOR T22[7];
   T13C_TRT_M1 : ALIAS FOR T22[7].PRE;
   T13C_TRT_M2 : ALIAS FOR T22[7].ACC;
   T13C_TRT_O : ALIAS FOR T22[5];
   T13C_TRT_O1 : ALIAS FOR T22[5].PRE;
   T13C_TRT_O2 : ALIAS FOR T22[5].ACC;
   T14_AIR_GT : ALIAS FOR I1.9;
   T14_AIR_SV : ALIAS FOR O9.9;
   T14_ASCII : ALIAS FOR B17[14].1;
   T14_ASSII : ALIAS FOR A16[142];
   T14_ASSII1 : ALIAS FOR A16[145];
   T14_AUTO_A : ALIAS FOR T4[64];
   T14_AUTO_A1 : ALIAS FOR T4[64].PRE;
   T14_AUTO_A2 : ALIAS FOR T4[64].ACC;
   T14_AUTO_M : ALIAS FOR B3[14].1;
   T14_AUTO_S : ALIAS FOR B3[14].14;
   T14_BINDIC : ALIAS FOR I4.14;
   T14_CAL_CL : ALIAS FOR B15[54].3;
   T14_CAL_LA : ALIAS FOR B15[54].2;
   T14_CAL_OP : ALIAS FOR B15[54].4;
   T14_CAL_ST : ALIAS FOR B15[54].1;
   T14_CLOSE : ALIAS FOR O9.10;
   T14_CLOSE1 : ALIAS FOR B3[14].9;
   T14_CLOSE2 : ALIAS FOR B3[14].11;
   T14_CORREC : ALIAS FOR F8[8];
   T14_DLY_TR : ALIAS FOR T4[6];
   T14_DLY_TR1 : ALIAS FOR T4[6].PRE;
   T14_DLY_TR2 : ALIAS FOR T4[6].ACC;
   T14_DLY_TR3 : ALIAS FOR T4[7];
   T14_DLY_TR4 : ALIAS FOR T4[7].PRE;
   T14_DLY_TR5 : ALIAS FOR T4[7].ACC;
   T14_FAULT : ALIAS FOR B3[14].15;
   T14_GATE_C : ALIAS FOR C5[14];
   T14_GATE_C1 : ALIAS FOR C5[14].PRE;
   T14_GATE_C2 : ALIAS FOR C5[14].ACC;
   T14_HOLD_A : ALIAS FOR B3[14].3;
   T14_HOLD_M : ALIAS FOR B3[14].6;
   T14_K_FACT : ALIAS FOR F8[7];
   T14_LOW_BI : ALIAS FOR B15[14].2;
   T14_MTR_GT : ALIAS FOR I1.11;
   T14_NO_PAS : ALIAS FOR B17[14].2;
   T14_NULL_V : ALIAS FOR A16[148];
   T14_NULL_V1 : ALIAS FOR A16[149];
   T14_OP_DEF : ALIAS FOR A16[146];
   T14_OP_DEF1 : ALIAS FOR A16[147];
   T14_OP_NAM : ALIAS FOR A16[143];
   T14_OP_NAM1 : ALIAS FOR A16[144];
   T14_OPEN_A : ALIAS FOR B3[14].8;
   T14_OPEN_M : ALIAS FOR O9.11;
   T14_OPEN_M1 : ALIAS FOR B3[14].10;
   T14_RELEAS : ALIAS FOR B3[14].5;
   T14_RESET : ALIAS FOR B3[14].7;
   T14_SET_AU : ALIAS FOR B3[14].2;
   T14_SET_DE : ALIAS FOR B3[2].3;
   T14_SET_LO : ALIAS FOR B3[14].13;
   T14_SET_MA : ALIAS FOR B3[14].12;
   T14_SET_NA : ALIAS FOR A16[140];
   T14_SET_NA1 : ALIAS FOR A16[141];
   T14_SET_NA2 : ALIAS FOR B17[14].0;
   T14_STOP_A : ALIAS FOR B3[14].4;
   T14_TREAT : ALIAS FOR B3[14].0;
   T14_TRT_MO : ALIAS FOR T4[44];
   T14_TRT_MO1 : ALIAS FOR T4[44].PRE;
   T14_TRT_MO2 : ALIAS FOR T4[44].ACC;
   T15_AIR_GT : ALIAS FOR I1.12;
   T15_AIR_SV : ALIAS FOR O9.12;
   T15_ASCII : ALIAS FOR B17[15].1;
   T15_ASSII : ALIAS FOR A16[152];
   T15_ASSII1 : ALIAS FOR A16[155];
   T15_AUTO_A : ALIAS FOR T4[65];
   T15_AUTO_A1 : ALIAS FOR T4[65].PRE;
   T15_AUTO_A2 : ALIAS FOR T4[65].ACC;
   T15_AUTO_M : ALIAS FOR B3[15].1;
   T15_AUTO_S : ALIAS FOR B3[15].14;
   T15_BINDIC : ALIAS FOR I4.15;
   T15_CAL_CL : ALIAS FOR B15[55].3;
   T15_CAL_LA : ALIAS FOR B15[55].2;
   T15_CAL_OP : ALIAS FOR B15[55].4;
   T15_CAL_ST : ALIAS FOR B15[55].1;
   T15_CLOSE : ALIAS FOR O9.13;
   T15_CLOSE1 : ALIAS FOR B3[15].9;
   T15_CLOSE2 : ALIAS FOR B3[15].11;
   T15_CORREC : ALIAS FOR F8[10];
   T15_FAULT : ALIAS FOR B3[15].15;
   T15_GATE_C : ALIAS FOR C5[15];
   T15_GATE_C1 : ALIAS FOR C5[15].PRE;
   T15_GATE_C2 : ALIAS FOR C5[15].ACC;
   T15_HOLD_A : ALIAS FOR B3[15].3;
   T15_HOLD_M : ALIAS FOR B3[15].6;
   T15_K_FACT : ALIAS FOR F8[9];
   T15_LOW_BI : ALIAS FOR B15[15].2;
   T15_MTR_GT : ALIAS FOR I1.14;
   T15_NO_PAS : ALIAS FOR B17[15].2;
   T15_NULL_V : ALIAS FOR A16[158];
   T15_NULL_V1 : ALIAS FOR A16[159];
   T15_OP_DEF : ALIAS FOR A16[156];
   T15_OP_DEF1 : ALIAS FOR A16[157];
   T15_OP_NAM : ALIAS FOR A16[153];
   T15_OP_NAM1 : ALIAS FOR A16[154];
   T15_OPEN_A : ALIAS FOR B3[15].8;
   T15_OPEN_M : ALIAS FOR O9.14;
   T15_OPEN_M1 : ALIAS FOR B3[15].10;
   T15_RELEAS : ALIAS FOR B3[15].5;
   T15_RESET : ALIAS FOR B3[15].7;
   T15_SET_AU : ALIAS FOR B3[15].2;
   T15_SET_DE : ALIAS FOR B3[2].4;
   T15_SET_LO : ALIAS FOR B3[15].13;
   T15_SET_MA : ALIAS FOR B3[15].12;
   T15_SET_NA : ALIAS FOR A16[150];
   T15_SET_NA1 : ALIAS FOR A16[151];
   T15_SET_NA2 : ALIAS FOR B17[15].0;
   T15_STOP_A : ALIAS FOR B3[15].4;
   T15_TREAT : ALIAS FOR B3[15].0;
   T15_TRT_MO : ALIAS FOR T4[45];
   T15_TRT_MO1 : ALIAS FOR T4[45].PRE;
   T15_TRT_MO2 : ALIAS FOR T4[45].ACC;
   T15_TRT_OF : ALIAS FOR T4[9];
   T15_TRT_OF1 : ALIAS FOR T4[9].PRE;
   T15_TRT_OF2 : ALIAS FOR T4[9].ACC;
   T15_TRT_ON : ALIAS FOR T4[8];
   T15_TRT_ON1 : ALIAS FOR T4[8].PRE;
   T15_TRT_ON2 : ALIAS FOR T4[8].ACC;
   T16_AIR_GA : ALIAS FOR I2.0;
   T16_AIR_SV : ALIAS FOR O10.0;
   T16_ASCII : ALIAS FOR B17[16].1;
   T16_ASSII : ALIAS FOR A16[162];
   T16_ASSII1 : ALIAS FOR A16[165];
   T16_AUTO_A : ALIAS FOR T4[66];
   T16_AUTO_A1 : ALIAS FOR T4[66].PRE;
   T16_AUTO_A2 : ALIAS FOR T4[66].ACC;
   T16_AUTO_M : ALIAS FOR B3[16].1;
   T16_AUTO_S : ALIAS FOR B3[16].14;
   T16_BINDIC : ALIAS FOR I4.9;
   T16_CAL_CL : ALIAS FOR B15[56].3;
   T16_CAL_LA : ALIAS FOR B15[56].2;
   T16_CAL_OP : ALIAS FOR B15[56].4;
   T16_CAL_ST : ALIAS FOR B15[56].1;
   T16_CLOSE : ALIAS FOR O10.1;
   T16_CLOSE1 : ALIAS FOR B3[16].9;
   T16_CLOSE2 : ALIAS FOR B3[16].11;
   T16_CORREC : ALIAS FOR F8[12];
   T16_FAULT : ALIAS FOR B3[16].15;
   T16_GATE_C : ALIAS FOR C5[16];
   T16_GATE_C1 : ALIAS FOR C5[16].PRE;
   T16_GATE_C2 : ALIAS FOR C5[16].ACC;
   T16_HOLD_A : ALIAS FOR B3[16].3;
   T16_HOLD_M : ALIAS FOR B3[16].6;
   T16_K_FACT : ALIAS FOR F8[11];
   T16_LOW_BI : ALIAS FOR B15[16].2;
   T16_METER : ALIAS FOR I2.2;
   T16_NO_PAS : ALIAS FOR B17[16].2;
   T16_NULL_V : ALIAS FOR A16[168];
   T16_NULL_V1 : ALIAS FOR A16[169];
   T16_OP_DEF : ALIAS FOR A16[166];
   T16_OP_DEF1 : ALIAS FOR A16[167];
   T16_OP_NAM : ALIAS FOR A16[163];
   T16_OP_NAM1 : ALIAS FOR A16[164];
   T16_OPEN_A : ALIAS FOR B3[16].8;
   T16_OPEN_M : ALIAS FOR O10.2;
   T16_OPEN_M1 : ALIAS FOR B3[16].10;
   T16_RELEAS : ALIAS FOR B3[16].5;
   T16_RESET : ALIAS FOR B3[16].7;
   T16_SET_AU : ALIAS FOR B3[16].2;
   T16_SET_DE : ALIAS FOR B3[2].5;
   T16_SET_LO : ALIAS FOR B3[16].13;
   T16_SET_MA : ALIAS FOR B3[16].12;
   T16_SET_NA : ALIAS FOR A16[160];
   T16_SET_NA1 : ALIAS FOR A16[161];
   T16_SET_NA2 : ALIAS FOR B17[16].0;
   T16_STOP_A : ALIAS FOR B3[16].4;
   T16_TREAT : ALIAS FOR B3[16].0;
   T16_TRT_MO : ALIAS FOR T4[46];
   T16_TRT_MO1 : ALIAS FOR T4[46].PRE;
   T16_TRT_MO2 : ALIAS FOR T4[46].ACC;
   T16_TRT_OF : ALIAS FOR T4[11];
   T16_TRT_OF1 : ALIAS FOR T4[11].PRE;
   T16_TRT_OF2 : ALIAS FOR T4[11].ACC;
   T16_TRT_ON : ALIAS FOR T4[10];
   T16_TRT_ON1 : ALIAS FOR T4[10].PRE;
   T16_TRT_ON2 : ALIAS FOR T4[10].ACC;
   T17_AIR_GA : ALIAS FOR I2.3;
   T17_AIR_SV : ALIAS FOR O10.3;
   T17_ASCII : ALIAS FOR B17[17].1;
   T17_ASSII : ALIAS FOR A16[172];
   T17_ASSII1 : ALIAS FOR A16[175];
   T17_AUTO_A : ALIAS FOR T4[67];
   T17_AUTO_A1 : ALIAS FOR T4[67].PRE;
   T17_AUTO_A2 : ALIAS FOR T4[67].ACC;
   T17_AUTO_M : ALIAS FOR B3[17].1;
   T17_AUTO_S : ALIAS FOR B3[17].14;
   T17_BINDIC : ALIAS FOR I4.10;
   T17_CAL_CL : ALIAS FOR B15[57].3;
   T17_CAL_LA : ALIAS FOR B15[57].2;
   T17_CAL_OP : ALIAS FOR B15[57].4;
   T17_CAL_ST : ALIAS FOR B15[57].1;
   T17_CLOSE : ALIAS FOR O10.4;
   T17_CLOSE1 : ALIAS FOR B3[17].9;
   T17_CLOSE2 : ALIAS FOR B3[17].11;
   T17_CORREC : ALIAS FOR F8[14];
   T17_FAULT : ALIAS FOR B3[17].15;
   T17_GATE_C : ALIAS FOR C5[17];
   T17_GATE_C1 : ALIAS FOR C5[17].PRE;
   T17_GATE_C2 : ALIAS FOR C5[17].ACC;
